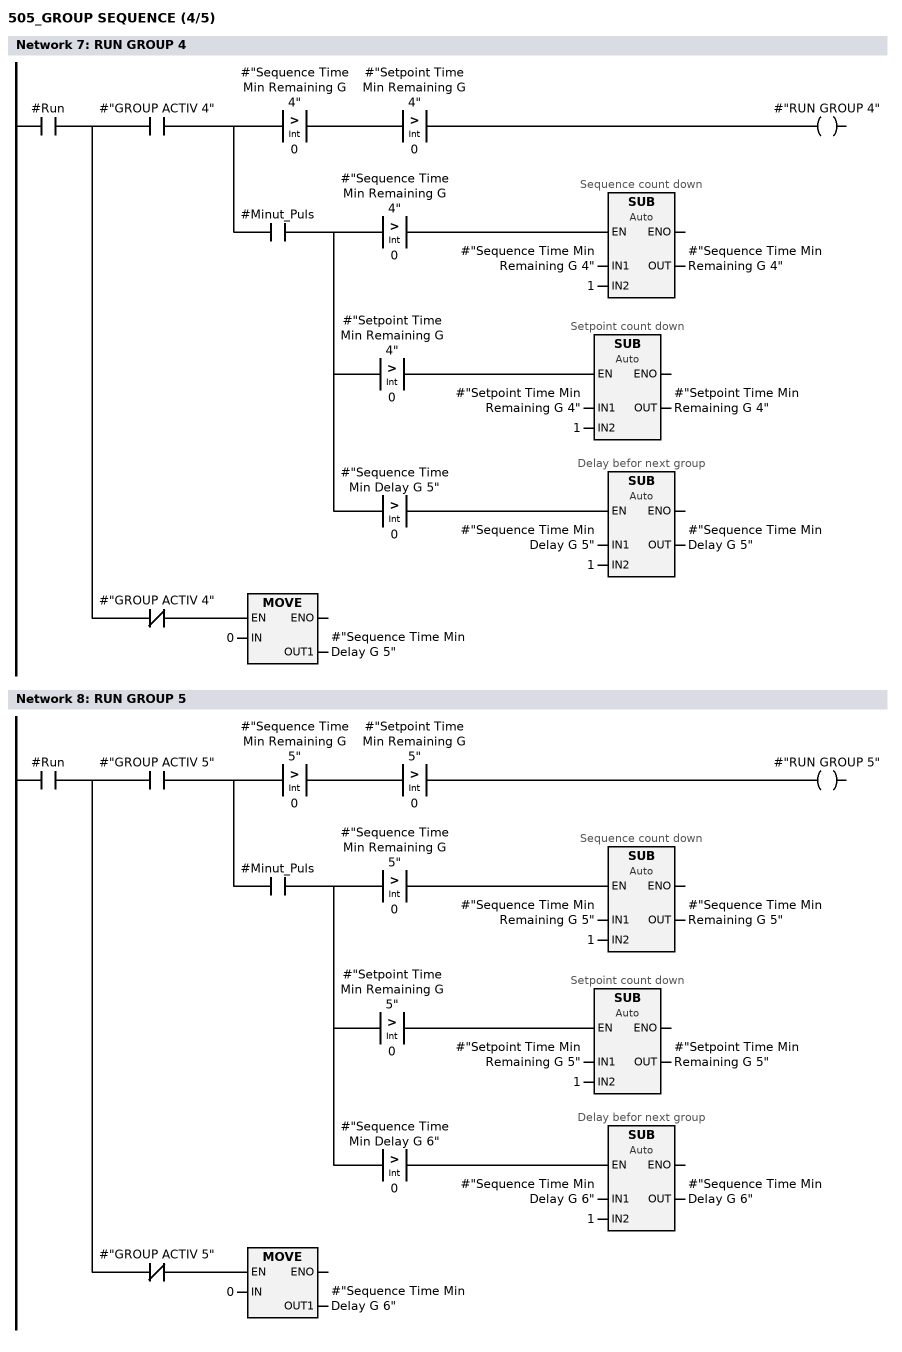
   RUNG wire#powerrail
      Contact( #Run )
      wire#w1
      Contact( #"GROUP ACTIV 4" )
      wire#w2
      { S7_Templates := "SrcType := Int" } GT_Contact(in1 := #"Sequence Time Min Remaining G 4", in2 := 0)
      { S7_Templates := "SrcType := Int" } GT_Contact(in1 := #"Setpoint Time Min Remaining G 4", in2 := 0)
      Coil( #"RUN GROUP 4" )
   END_RUNG
   RUNG wire#w2
      Contact( #Minut_Puls )
      wire#w3
      { S7_Templates := "SrcType := Int" } GT_Contact(in1 := #"Sequence Time Min Remaining G 4", in2 := 0)
      Sub(in1 := #"Sequence Time Min Remaining G 4", in2 := 1, out => #"Sequence Time Min Remaining G 4")   // Sequence count down
   END_RUNG
   RUNG wire#w3
      { S7_Templates := "SrcType := Int" } GT_Contact(in1 := #"Setpoint Time Min Remaining G 4", in2 := 0)
      Sub(in1 := #"Setpoint Time Min Remaining G 4", in2 := 1, out => #"Setpoint Time Min Remaining G 4")   // Setpoint count down
   END_RUNG
   RUNG wire#w3
      { S7_Templates := "SrcType := Int" } GT_Contact(in1 := #"Sequence Time Min Delay G 5", in2 := 0)
      Sub(in1 := #"Sequence Time Min Delay G 5", in2 := 1, out => #"Sequence Time Min Delay G 5")   // Delay befor next group
   END_RUNG
   RUNG wire#w1
      I_Contact( #"GROUP ACTIV 4" )
      Move(in := 0, out1 => #"Sequence Time Min Delay G 5")
   END_RUNG
   // the same network as SCL:
   #_w1 := #Run AND #"GROUP ACTIV 4";
   #"RUN GROUP 4" := #_w1 AND (#"Sequence Time Min Remaining G 4" > 0) AND (#"Setpoint Time Min Remaining G 4" > 0);
   #_w2 := #_w1 AND #Minut_Puls;
   IF #_w2 AND (#"Sequence Time Min Remaining G 4" > 0) THEN
       #"Sequence Time Min Remaining G 4" := #"Sequence Time Min Remaining G 4" - 1;   // Sequence count down
   END_IF;
   IF #_w2 AND (#"Setpoint Time Min Remaining G 4" > 0) THEN
       #"Setpoint Time Min Remaining G 4" := #"Setpoint Time Min Remaining G 4" - 1;   // Setpoint count down
   END_IF;
   IF #_w2 AND (#"Sequence Time Min Delay G 5" > 0) THEN
       #"Sequence Time Min Delay G 5" := #"Sequence Time Min Delay G 5" - 1;   // Delay befor next group
   END_IF;
   IF #Run AND NOT #"GROUP ACTIV 4" THEN #"Sequence Time Min Delay G 5" := 0; END_IF;
END_REGION

REGION Network 8: RUN GROUP 5
   RUNG wire#powerrail
      Contact( #Run )
      wire#w1
      Contact( #"GROUP ACTIV 5" )
      wire#w2
      { S7_Templates := "SrcType := Int" } GT_Contact(in1 := #"Sequence Time Min Remaining G 5", in2 := 0)
      { S7_Templates := "SrcType := Int" } GT_Contact(in1 := #"Setpoint Time Min Remaining G 5", in2 := 0)
      Coil( #"RUN GROUP 5" )
   END_RUNG
   RUNG wire#w2
      Contact( #Minut_Puls )
      wire#w3
      { S7_Templates := "SrcType := Int" } GT_Contact(in1 := #"Sequence Time Min Remaining G 5", in2 := 0)
      Sub(in1 := #"Sequence Time Min Remaining G 5", in2 := 1, out => #"Sequence Time Min Remaining G 5")   // Sequence count down
   END_RUNG
   RUNG wire#w3
      { S7_Templates := "SrcType := Int" } GT_Contact(in1 := #"Setpoint Time Min Remaining G 5", in2 := 0)
      Sub(in1 := #"Setpoint Time Min Remaining G 5", in2 := 1, out => #"Setpoint Time Min Remaining G 5")   // Setpoint count down
   END_RUNG
   RUNG wire#w3
      { S7_Templates := "SrcType := Int" } GT_Contact(in1 := #"Sequence Time Min Delay G 6", in2 := 0)
      Sub(in1 := #"Sequence Time Min Delay G 6", in2 := 1, out => #"Sequence Time Min Delay G 6")   // Delay befor next group
   END_RUNG
   RUNG wire#w1
      I_Contact( #"GROUP ACTIV 5" )
      Move(in := 0, out1 => #"Sequence Time Min Delay G 6")
   END_RUNG
   // the same network as SCL:
   #_w1 := #Run AND #"GROUP ACTIV 5";
   #"RUN GROUP 5" := #_w1 AND (#"Sequence Time Min Remaining G 5" > 0) AND (#"Setpoint Time Min Remaining G 5" > 0);
   #_w2 := #_w1 AND #Minut_Puls;
   IF #_w2 AND (#"Sequence Time Min Remaining G 5" > 0) THEN
       #"Sequence Time Min Remaining G 5" := #"Sequence Time Min Remaining G 5" - 1;   // Sequence count down
   END_IF;
   IF #_w2 AND (#"Setpoint Time Min Remaining G 5" > 0) THEN
       #"Setpoint Time Min Remaining G 5" := #"Setpoint Time Min Remaining G 5" - 1;   // Setpoint count down
   END_IF;
   IF #_w2 AND (#"Sequence Time Min Delay G 6" > 0) THEN
       #"Sequence Time Min Delay G 6" := #"Sequence Time Min Delay G 6" - 1;   // Delay befor next group
   END_IF;
   IF #Run AND NOT #"GROUP ACTIV 5" THEN #"Sequence Time Min Delay G 6" := 0; END_IF;
END_REGION

REGION Network 9: RUN GROUP 6
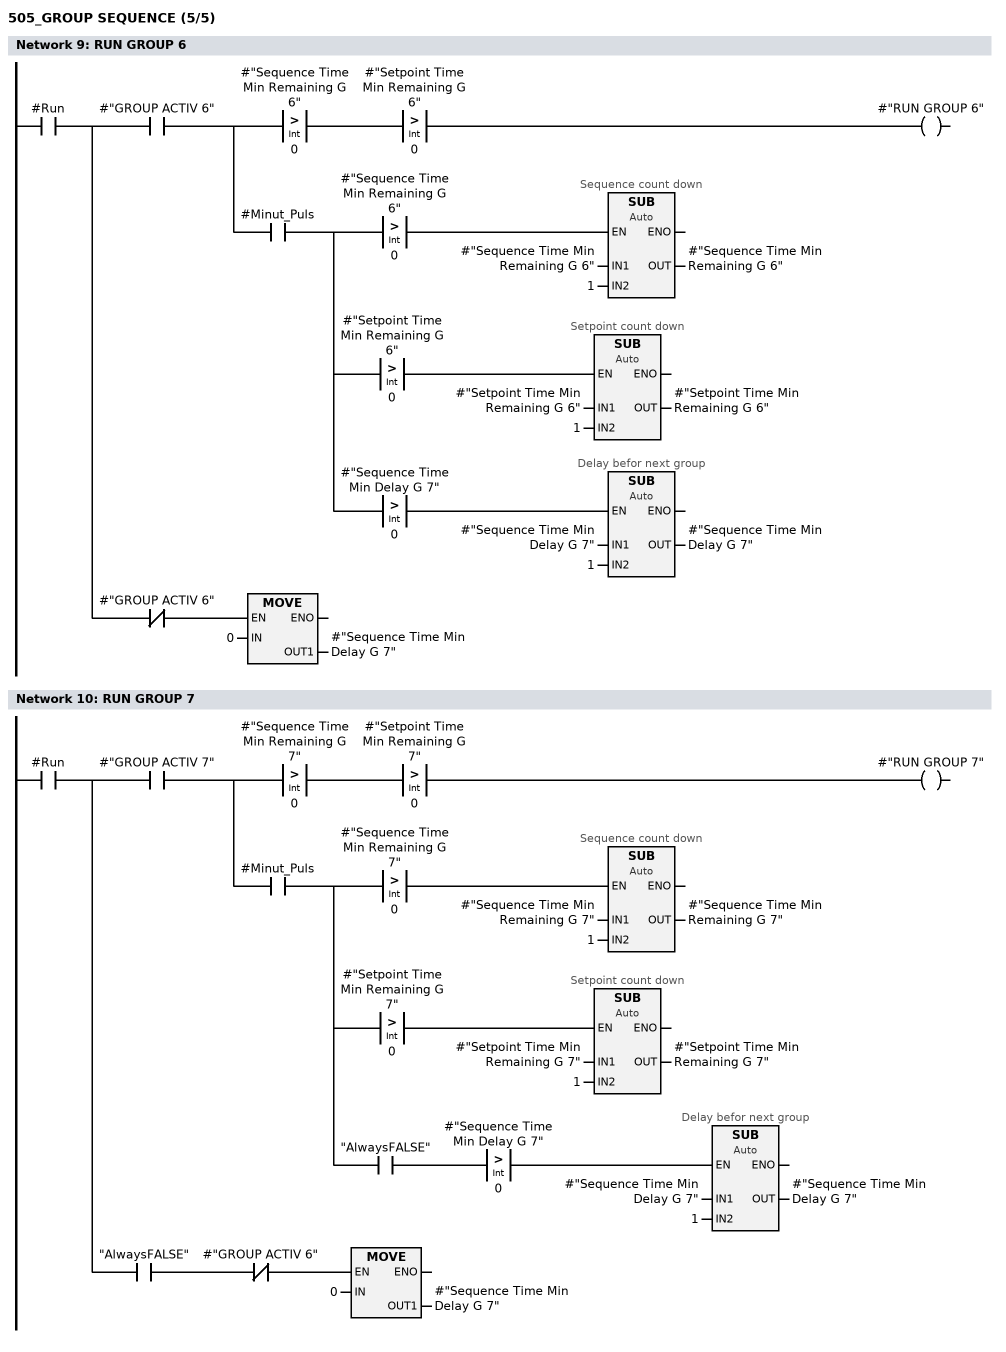
   RUNG wire#powerrail
      Contact( #Run )
      wire#w1
      Contact( #"GROUP ACTIV 6" )
      wire#w2
      { S7_Templates := "SrcType := Int" } GT_Contact(in1 := #"Sequence Time Min Remaining G 6", in2 := 0)
      { S7_Templates := "SrcType := Int" } GT_Contact(in1 := #"Setpoint Time Min Remaining G 6", in2 := 0)
      Coil( #"RUN GROUP 6" )
   END_RUNG
   RUNG wire#w2
      Contact( #Minut_Puls )
      wire#w3
      { S7_Templates := "SrcType := Int" } GT_Contact(in1 := #"Sequence Time Min Remaining G 6", in2 := 0)
      Sub(in1 := #"Sequence Time Min Remaining G 6", in2 := 1, out => #"Sequence Time Min Remaining G 6")   // Sequence count down
   END_RUNG
   RUNG wire#w3
      { S7_Templates := "SrcType := Int" } GT_Contact(in1 := #"Setpoint Time Min Remaining G 6", in2 := 0)
      Sub(in1 := #"Setpoint Time Min Remaining G 6", in2 := 1, out => #"Setpoint Time Min Remaining G 6")   // Setpoint count down
   END_RUNG
   RUNG wire#w3
      { S7_Templates := "SrcType := Int" } GT_Contact(in1 := #"Sequence Time Min Delay G 7", in2 := 0)
      Sub(in1 := #"Sequence Time Min Delay G 7", in2 := 1, out => #"Sequence Time Min Delay G 7")   // Delay befor next group
   END_RUNG
   RUNG wire#w1
      I_Contact( #"GROUP ACTIV 6" )
      Move(in := 0, out1 => #"Sequence Time Min Delay G 7")
   END_RUNG
   // the same network as SCL:
   #_w1 := #Run AND #"GROUP ACTIV 6";
   #"RUN GROUP 6" := #_w1 AND (#"Sequence Time Min Remaining G 6" > 0) AND (#"Setpoint Time Min Remaining G 6" > 0);
   #_w2 := #_w1 AND #Minut_Puls;
   IF #_w2 AND (#"Sequence Time Min Remaining G 6" > 0) THEN
       #"Sequence Time Min Remaining G 6" := #"Sequence Time Min Remaining G 6" - 1;   // Sequence count down
   END_IF;
   IF #_w2 AND (#"Setpoint Time Min Remaining G 6" > 0) THEN
       #"Setpoint Time Min Remaining G 6" := #"Setpoint Time Min Remaining G 6" - 1;   // Setpoint count down
   END_IF;
   IF #_w2 AND (#"Sequence Time Min Delay G 7" > 0) THEN
       #"Sequence Time Min Delay G 7" := #"Sequence Time Min Delay G 7" - 1;   // Delay befor next group
   END_IF;
   IF #Run AND NOT #"GROUP ACTIV 6" THEN #"Sequence Time Min Delay G 7" := 0; END_IF;
END_REGION

REGION Network 10: RUN GROUP 7
   RUNG wire#powerrail
      Contact( #Run )
      wire#w1
      Contact( #"GROUP ACTIV 7" )
      wire#w2
      { S7_Templates := "SrcType := Int" } GT_Contact(in1 := #"Sequence Time Min Remaining G 7", in2 := 0)
      { S7_Templates := "SrcType := Int" } GT_Contact(in1 := #"Setpoint Time Min Remaining G 7", in2 := 0)
      Coil( #"RUN GROUP 7" )
   END_RUNG
   RUNG wire#w2
      Contact( #Minut_Puls )
      wire#w3
      { S7_Templates := "SrcType := Int" } GT_Contact(in1 := #"Sequence Time Min Remaining G 7", in2 := 0)
      Sub(in1 := #"Sequence Time Min Remaining G 7", in2 := 1, out => #"Sequence Time Min Remaining G 7")   // Sequence count down
   END_RUNG
   RUNG wire#w3
      { S7_Templates := "SrcType := Int" } GT_Contact(in1 := #"Setpoint Time Min Remaining G 7", in2 := 0)
      Sub(in1 := #"Setpoint Time Min Remaining G 7", in2 := 1, out => #"Setpoint Time Min Remaining G 7")   // Setpoint count down
   END_RUNG
   RUNG wire#w3
      Contact( "AlwaysFALSE" )
      { S7_Templates := "SrcType := Int" } GT_Contact(in1 := #"Sequence Time Min Delay G 7", in2 := 0)
      Sub(in1 := #"Sequence Time Min Delay G 7", in2 := 1, out => #"Sequence Time Min Delay G 7")   // Delay befor next group
   END_RUNG
   RUNG wire#w1
      Contact( "AlwaysFALSE" )
      I_Contact( #"GROUP ACTIV 6" )
      Move(in := 0, out1 => #"Sequence Time Min Delay G 7")
   END_RUNG
   // the same network as SCL:
   #_w1 := #Run AND #"GROUP ACTIV 7";
   #"RUN GROUP 7" := #_w1 AND (#"Sequence Time Min Remaining G 7" > 0) AND (#"Setpoint Time Min Remaining G 7" > 0);
   #_w2 := #_w1 AND #Minut_Puls;
   IF #_w2 AND (#"Sequence Time Min Remaining G 7" > 0) THEN
       #"Sequence Time Min Remaining G 7" := #"Sequence Time Min Remaining G 7" - 1;   // Sequence count down
   END_IF;
   IF #_w2 AND (#"Setpoint Time Min Remaining G 7" > 0) THEN
       #"Setpoint Time Min Remaining G 7" := #"Setpoint Time Min Remaining G 7" - 1;   // Setpoint count down
   END_IF;
   IF #_w2 AND "AlwaysFALSE" AND (#"Sequence Time Min Delay G 7" > 0) THEN
       #"Sequence Time Min Delay G 7" := #"Sequence Time Min Delay G 7" - 1;   // Delay befor next group
   END_IF;
   IF #Run AND "AlwaysFALSE" AND NOT #"GROUP ACTIV 6" THEN #"Sequence Time Min Delay G 7" := 0; END_IF;
END_REGION
END_FUNCTION_BLOCK

FUNCTION_BLOCK "Binary Imputs ADD"   // FB506, LAD
{ S7_Optimized_Access := 'TRUE' }
VERSION : 0.1
   VAR_INPUT
      "BI 1" : Bool;
      "BI 2" : Bool;
      "BI 3" : Bool;
      "BI 4" : Bool;
      "BI 5" : Bool;
      "BI 6" : Bool;
      "BI 7" : Bool;
      "BI 8" : Bool;
      "BI 9" : Bool;
      "BI 10" : Bool;
      "BI 11" : Bool;
      "BI 12" : Bool;
      "BI 13" : Bool;
      "BI 14" : Bool;
      "BI 15" : Bool;
      "BI 16" : Bool;
      "BI 17" : Bool;
      "BI 18" : Bool;
      "BI 19" : Bool;
      "BI 20" : Bool;
      "BI 21" : Bool;
      "BI 22" : Bool;
      "BI 23" : Bool;
      "BI 24" : Bool;
   END_VAR
   VAR_OUTPUT
      "BI Number" : Int;
   END_VAR
   VAR
      "BI Interm 1" : Int;
      "BI Interm 2" : Int;
      "BI Interm 3" : Int;
      "BI Interm 4" : Int;
      "BI Interm 5" : Int;
      "BI Interm 6" : Int;
      "BI Interm 7" : Int;
      "BI Interm 8" : Int;
      "BI Interm 9" : Int;
      "BI Interm 10" : Int;
      "BI Interm 11" : Int;
      "BI Interm 12" : Int;
      "BI Interm 13" : Int;
      "BI Interm 14" : Int;
      "BI Interm 15" : Int;
      "BI Interm 16" : Int;
      "BI Interm 17" : Int;
      "BI Interm 18" : Int;
      "BI Interm 19" : Int;
      "BI Interm 20" : Int;
      "BI Interm 21" : Int;
      "BI Interm 22" : Int;
      "BI Interm 23" : Int;
      "BI Interm 24" : Int;
   END_VAR
BEGIN

REGION Network 1: 1
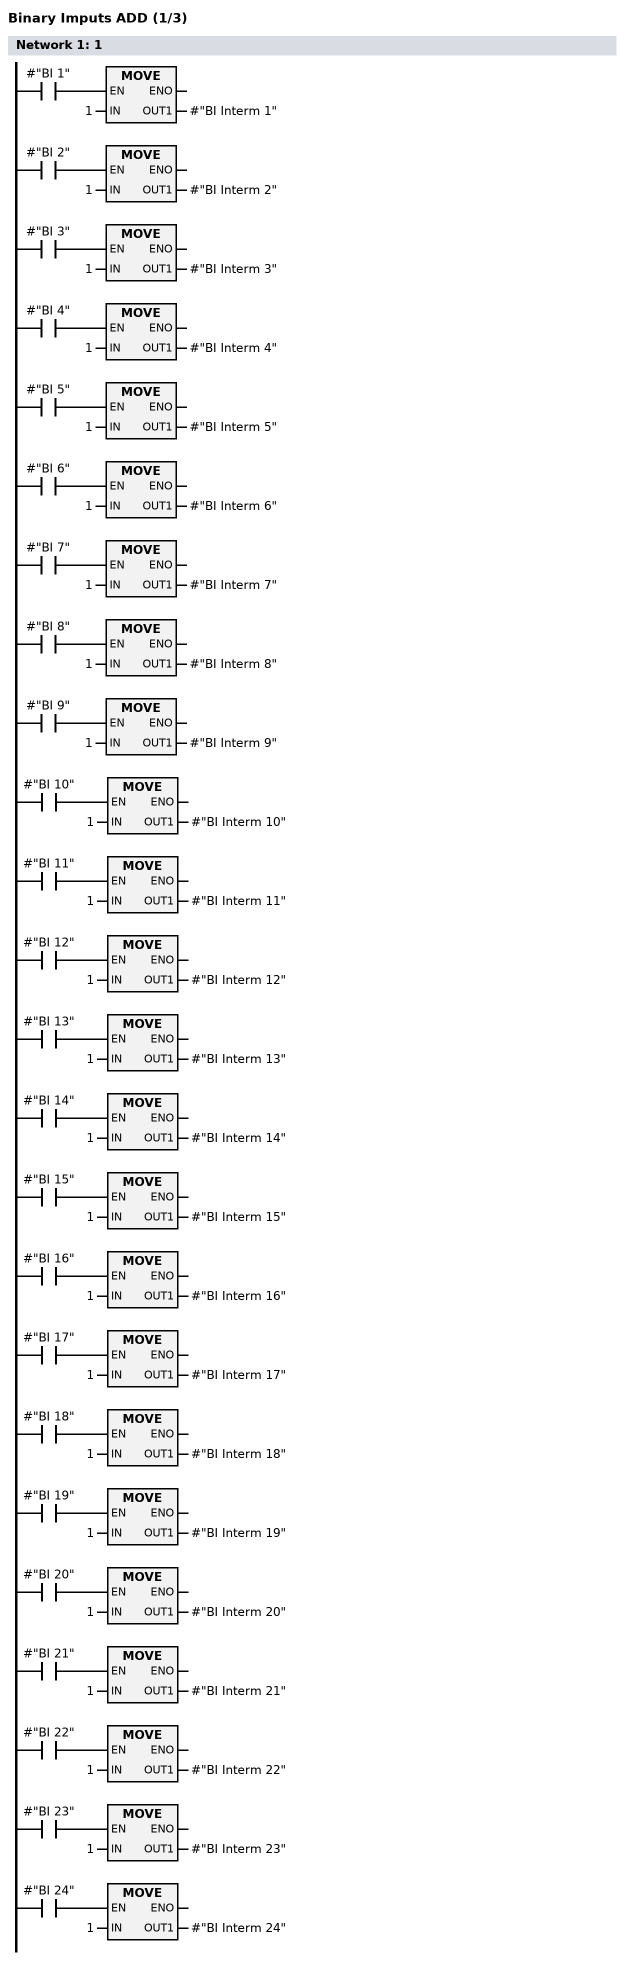
   RUNG wire#powerrail
      Contact( #"BI 1" )
      Move(in := 1, out1 => #"BI Interm 1")
   END_RUNG
   RUNG wire#powerrail
      Contact( #"BI 2" )
      Move(in := 1, out1 => #"BI Interm 2")
   END_RUNG
   RUNG wire#powerrail
      Contact( #"BI 3" )
      Move(in := 1, out1 => #"BI Interm 3")
   END_RUNG
   RUNG wire#powerrail
      Contact( #"BI 4" )
      Move(in := 1, out1 => #"BI Interm 4")
   END_RUNG
   RUNG wire#powerrail
      Contact( #"BI 5" )
      Move(in := 1, out1 => #"BI Interm 5")
   END_RUNG
   RUNG wire#powerrail
      Contact( #"BI 6" )
      Move(in := 1, out1 => #"BI Interm 6")
   END_RUNG
   RUNG wire#powerrail
      Contact( #"BI 7" )
      Move(in := 1, out1 => #"BI Interm 7")
   END_RUNG
   RUNG wire#powerrail
      Contact( #"BI 8" )
      Move(in := 1, out1 => #"BI Interm 8")
   END_RUNG
   RUNG wire#powerrail
      Contact( #"BI 9" )
      Move(in := 1, out1 => #"BI Interm 9")
   END_RUNG
   RUNG wire#powerrail
      Contact( #"BI 10" )
      Move(in := 1, out1 => #"BI Interm 10")
   END_RUNG
   RUNG wire#powerrail
      Contact( #"BI 11" )
      Move(in := 1, out1 => #"BI Interm 11")
   END_RUNG
   RUNG wire#powerrail
      Contact( #"BI 12" )
      Move(in := 1, out1 => #"BI Interm 12")
   END_RUNG
   RUNG wire#powerrail
      Contact( #"BI 13" )
      Move(in := 1, out1 => #"BI Interm 13")
   END_RUNG
   RUNG wire#powerrail
      Contact( #"BI 14" )
      Move(in := 1, out1 => #"BI Interm 14")
   END_RUNG
   RUNG wire#powerrail
      Contact( #"BI 15" )
      Move(in := 1, out1 => #"BI Interm 15")
   END_RUNG
   RUNG wire#powerrail
      Contact( #"BI 16" )
      Move(in := 1, out1 => #"BI Interm 16")
   END_RUNG
   RUNG wire#powerrail
      Contact( #"BI 17" )
      Move(in := 1, out1 => #"BI Interm 17")
   END_RUNG
   RUNG wire#powerrail
      Contact( #"BI 18" )
      Move(in := 1, out1 => #"BI Interm 18")
   END_RUNG
   RUNG wire#powerrail
      Contact( #"BI 19" )
      Move(in := 1, out1 => #"BI Interm 19")
   END_RUNG
   RUNG wire#powerrail
      Contact( #"BI 20" )
      Move(in := 1, out1 => #"BI Interm 20")
   END_RUNG
   RUNG wire#powerrail
      Contact( #"BI 21" )
      Move(in := 1, out1 => #"BI Interm 21")
   END_RUNG
   RUNG wire#powerrail
      Contact( #"BI 22" )
      Move(in := 1, out1 => #"BI Interm 22")
   END_RUNG
   RUNG wire#powerrail
      Contact( #"BI 23" )
      Move(in := 1, out1 => #"BI Interm 23")
   END_RUNG
   RUNG wire#powerrail
      Contact( #"BI 24" )
      Move(in := 1, out1 => #"BI Interm 24")
   END_RUNG
   // the same network as SCL:
   IF #"BI 1" THEN #"BI Interm 1" := 1; END_IF;
   IF #"BI 2" THEN #"BI Interm 2" := 1; END_IF;
   IF #"BI 3" THEN #"BI Interm 3" := 1; END_IF;
   IF #"BI 4" THEN #"BI Interm 4" := 1; END_IF;
   IF #"BI 5" THEN #"BI Interm 5" := 1; END_IF;
   IF #"BI 6" THEN #"BI Interm 6" := 1; END_IF;
   IF #"BI 7" THEN #"BI Interm 7" := 1; END_IF;
   IF #"BI 8" THEN #"BI Interm 8" := 1; END_IF;
   IF #"BI 9" THEN #"BI Interm 9" := 1; END_IF;
   IF #"BI 10" THEN #"BI Interm 10" := 1; END_IF;
   IF #"BI 11" THEN #"BI Interm 11" := 1; END_IF;
   IF #"BI 12" THEN #"BI Interm 12" := 1; END_IF;
   IF #"BI 13" THEN #"BI Interm 13" := 1; END_IF;
   IF #"BI 14" THEN #"BI Interm 14" := 1; END_IF;
   IF #"BI 15" THEN #"BI Interm 15" := 1; END_IF;
   IF #"BI 16" THEN #"BI Interm 16" := 1; END_IF;
   IF #"BI 17" THEN #"BI Interm 17" := 1; END_IF;
   IF #"BI 18" THEN #"BI Interm 18" := 1; END_IF;
   IF #"BI 19" THEN #"BI Interm 19" := 1; END_IF;
   IF #"BI 20" THEN #"BI Interm 20" := 1; END_IF;
   IF #"BI 21" THEN #"BI Interm 21" := 1; END_IF;
   IF #"BI 22" THEN #"BI Interm 22" := 1; END_IF;
   IF #"BI 23" THEN #"BI Interm 23" := 1; END_IF;
   IF #"BI 24" THEN #"BI Interm 24" := 1; END_IF;
END_REGION

REGION Network 2: 0
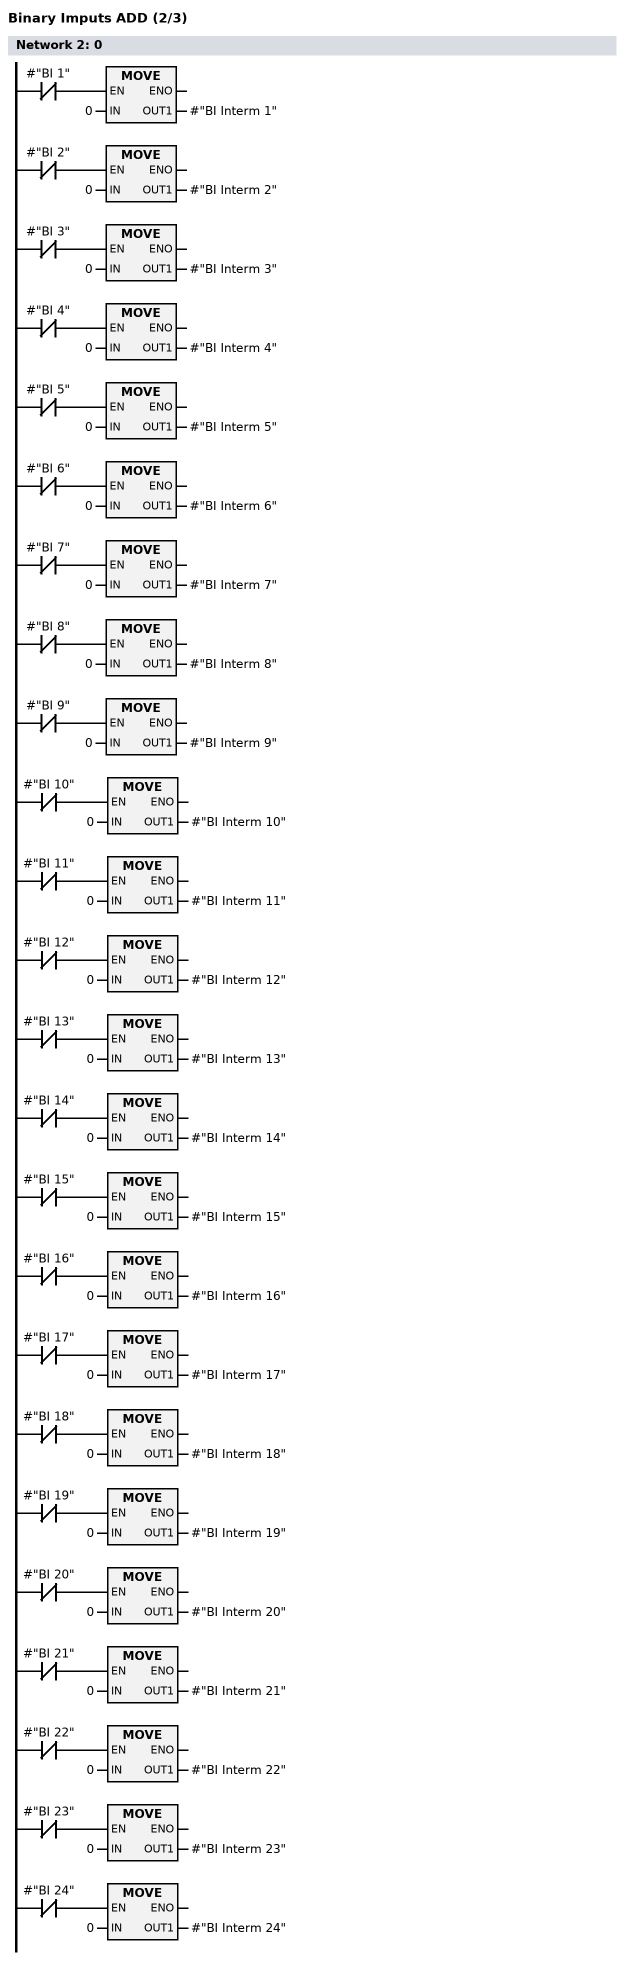
   RUNG wire#powerrail
      I_Contact( #"BI 1" )
      Move(in := 0, out1 => #"BI Interm 1")
   END_RUNG
   RUNG wire#powerrail
      I_Contact( #"BI 2" )
      Move(in := 0, out1 => #"BI Interm 2")
   END_RUNG
   RUNG wire#powerrail
      I_Contact( #"BI 3" )
      Move(in := 0, out1 => #"BI Interm 3")
   END_RUNG
   RUNG wire#powerrail
      I_Contact( #"BI 4" )
      Move(in := 0, out1 => #"BI Interm 4")
   END_RUNG
   RUNG wire#powerrail
      I_Contact( #"BI 5" )
      Move(in := 0, out1 => #"BI Interm 5")
   END_RUNG
   RUNG wire#powerrail
      I_Contact( #"BI 6" )
      Move(in := 0, out1 => #"BI Interm 6")
   END_RUNG
   RUNG wire#powerrail
      I_Contact( #"BI 7" )
      Move(in := 0, out1 => #"BI Interm 7")
   END_RUNG
   RUNG wire#powerrail
      I_Contact( #"BI 8" )
      Move(in := 0, out1 => #"BI Interm 8")
   END_RUNG
   RUNG wire#powerrail
      I_Contact( #"BI 9" )
      Move(in := 0, out1 => #"BI Interm 9")
   END_RUNG
   RUNG wire#powerrail
      I_Contact( #"BI 10" )
      Move(in := 0, out1 => #"BI Interm 10")
   END_RUNG
   RUNG wire#powerrail
      I_Contact( #"BI 11" )
      Move(in := 0, out1 => #"BI Interm 11")
   END_RUNG
   RUNG wire#powerrail
      I_Contact( #"BI 12" )
      Move(in := 0, out1 => #"BI Interm 12")
   END_RUNG
   RUNG wire#powerrail
      I_Contact( #"BI 13" )
      Move(in := 0, out1 => #"BI Interm 13")
   END_RUNG
   RUNG wire#powerrail
      I_Contact( #"BI 14" )
      Move(in := 0, out1 => #"BI Interm 14")
   END_RUNG
   RUNG wire#powerrail
      I_Contact( #"BI 15" )
      Move(in := 0, out1 => #"BI Interm 15")
   END_RUNG
   RUNG wire#powerrail
      I_Contact( #"BI 16" )
      Move(in := 0, out1 => #"BI Interm 16")
   END_RUNG
   RUNG wire#powerrail
      I_Contact( #"BI 17" )
      Move(in := 0, out1 => #"BI Interm 17")
   END_RUNG
   RUNG wire#powerrail
      I_Contact( #"BI 18" )
      Move(in := 0, out1 => #"BI Interm 18")
   END_RUNG
   RUNG wire#powerrail
      I_Contact( #"BI 19" )
      Move(in := 0, out1 => #"BI Interm 19")
   END_RUNG
   RUNG wire#powerrail
      I_Contact( #"BI 20" )
      Move(in := 0, out1 => #"BI Interm 20")
   END_RUNG
   RUNG wire#powerrail
      I_Contact( #"BI 21" )
      Move(in := 0, out1 => #"BI Interm 21")
   END_RUNG
   RUNG wire#powerrail
      I_Contact( #"BI 22" )
      Move(in := 0, out1 => #"BI Interm 22")
   END_RUNG
   RUNG wire#powerrail
      I_Contact( #"BI 23" )
      Move(in := 0, out1 => #"BI Interm 23")
   END_RUNG
   RUNG wire#powerrail
      I_Contact( #"BI 24" )
      Move(in := 0, out1 => #"BI Interm 24")
   END_RUNG
   // the same network as SCL:
   IF NOT #"BI 1" THEN #"BI Interm 1" := 0; END_IF;
   IF NOT #"BI 2" THEN #"BI Interm 2" := 0; END_IF;
   IF NOT #"BI 3" THEN #"BI Interm 3" := 0; END_IF;
   IF NOT #"BI 4" THEN #"BI Interm 4" := 0; END_IF;
   IF NOT #"BI 5" THEN #"BI Interm 5" := 0; END_IF;
   IF NOT #"BI 6" THEN #"BI Interm 6" := 0; END_IF;
   IF NOT #"BI 7" THEN #"BI Interm 7" := 0; END_IF;
   IF NOT #"BI 8" THEN #"BI Interm 8" := 0; END_IF;
   IF NOT #"BI 9" THEN #"BI Interm 9" := 0; END_IF;
   IF NOT #"BI 10" THEN #"BI Interm 10" := 0; END_IF;
   IF NOT #"BI 11" THEN #"BI Interm 11" := 0; END_IF;
   IF NOT #"BI 12" THEN #"BI Interm 12" := 0; END_IF;
   IF NOT #"BI 13" THEN #"BI Interm 13" := 0; END_IF;
   IF NOT #"BI 14" THEN #"BI Interm 14" := 0; END_IF;
   IF NOT #"BI 15" THEN #"BI Interm 15" := 0; END_IF;
   IF NOT #"BI 16" THEN #"BI Interm 16" := 0; END_IF;
   IF NOT #"BI 17" THEN #"BI Interm 17" := 0; END_IF;
   IF NOT #"BI 18" THEN #"BI Interm 18" := 0; END_IF;
   IF NOT #"BI 19" THEN #"BI Interm 19" := 0; END_IF;
   IF NOT #"BI 20" THEN #"BI Interm 20" := 0; END_IF;
   IF NOT #"BI 21" THEN #"BI Interm 21" := 0; END_IF;
   IF NOT #"BI 22" THEN #"BI Interm 22" := 0; END_IF;
   IF NOT #"BI 23" THEN #"BI Interm 23" := 0; END_IF;
   IF NOT #"BI 24" THEN #"BI Interm 24" := 0; END_IF;
END_REGION

REGION Network 3: ADD
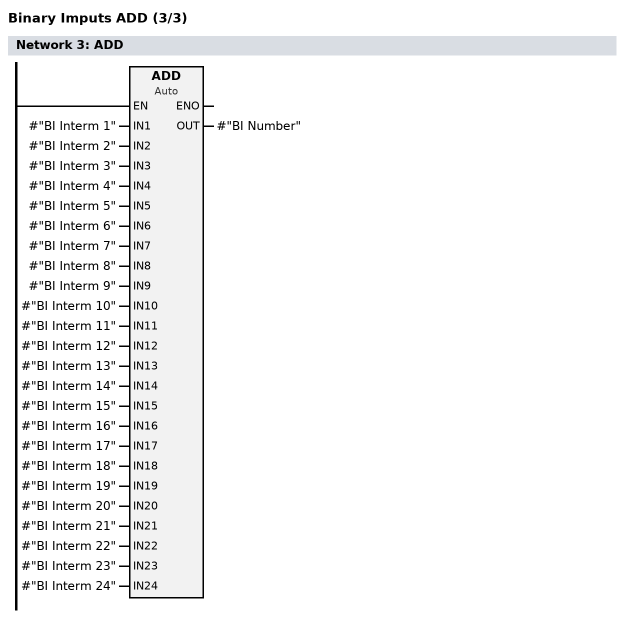
   RUNG wire#powerrail
      Add(in1 := #"BI Interm 1", in2 := #"BI Interm 2", in3 := #"BI Interm 3", in4 := #"BI Interm 4", in5 := #"BI Interm 5", in6 := #"BI Interm 6", in7 := #"BI Interm 7", in8 := #"BI Interm 8", in9 := #"BI Interm 9", in10 := #"BI Interm 10", in11 := #"BI Interm 11", in12 := #"BI Interm 12", in13 := #"BI Interm 13", in14 := #"BI Interm 14", in15 := #"BI Interm 15", in16 := #"BI Interm 16", in17 := #"BI Interm 17", in18 := #"BI Interm 18", in19 := #"BI Interm 19", in20 := #"BI Interm 20", in21 := #"BI Interm 21", in22 := #"BI Interm 22", in23 := #"BI Interm 23", in24 := #"BI Interm 24", out => #"BI Number")
   END_RUNG
   // the same network as SCL:
   #"BI Number" := #"BI Interm 1" + #"BI Interm 2" + #"BI Interm 3" + #"BI Interm 4" + #"BI Interm 5" + #"BI Interm 6" + #"BI Interm 7" + #"BI Interm 8" + #"BI Interm 9" + #"BI Interm 10" + #"BI Interm 11" + #"BI Interm 12" + #"BI Interm 13" + #"BI Interm 14" + #"BI Interm 15" + #"BI Interm 16" + #"BI Interm 17" + #"BI Interm 18" + #"BI Interm 19" + #"BI Interm 20" + #"BI Interm 21" + #"BI Interm 22" + #"BI Interm 23" + #"BI Interm 24";
END_REGION
END_FUNCTION_BLOCK

FUNCTION_BLOCK "HMI Indication Logic"   // FB507, LAD
{ S7_Optimized_Access := 'TRUE' }
VERSION : 0.1
   VAR_OUTPUT
      "FA Mode Selected" : Bool;
      "Tank Selected" : Bool;
      "Sequence Finished" : Bool;
   END_VAR
   VAR
      IEC_Timer_0_Instance : TON_TIME;
   END_VAR
BEGIN

REGION Network 1: FA Mode Selected
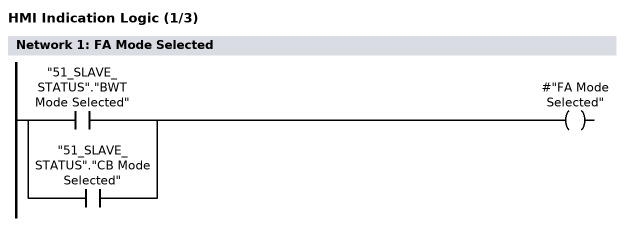
   RUNG wire#powerrail
      Contact( "51_SLAVE_STATUS"."BWT Mode Selected" )
      wire#w1
      Coil( #"FA Mode Selected" )
   END_RUNG
   RUNG wire#powerrail
      Contact( "51_SLAVE_STATUS"."CB Mode Selected" )
   END_RUNG wire#w1
   // the same network as SCL:
   #"FA Mode Selected" := "51_SLAVE_STATUS"."BWT Mode Selected" OR "51_SLAVE_STATUS"."CB Mode Selected";
END_REGION

REGION Network 2: Tank Selected
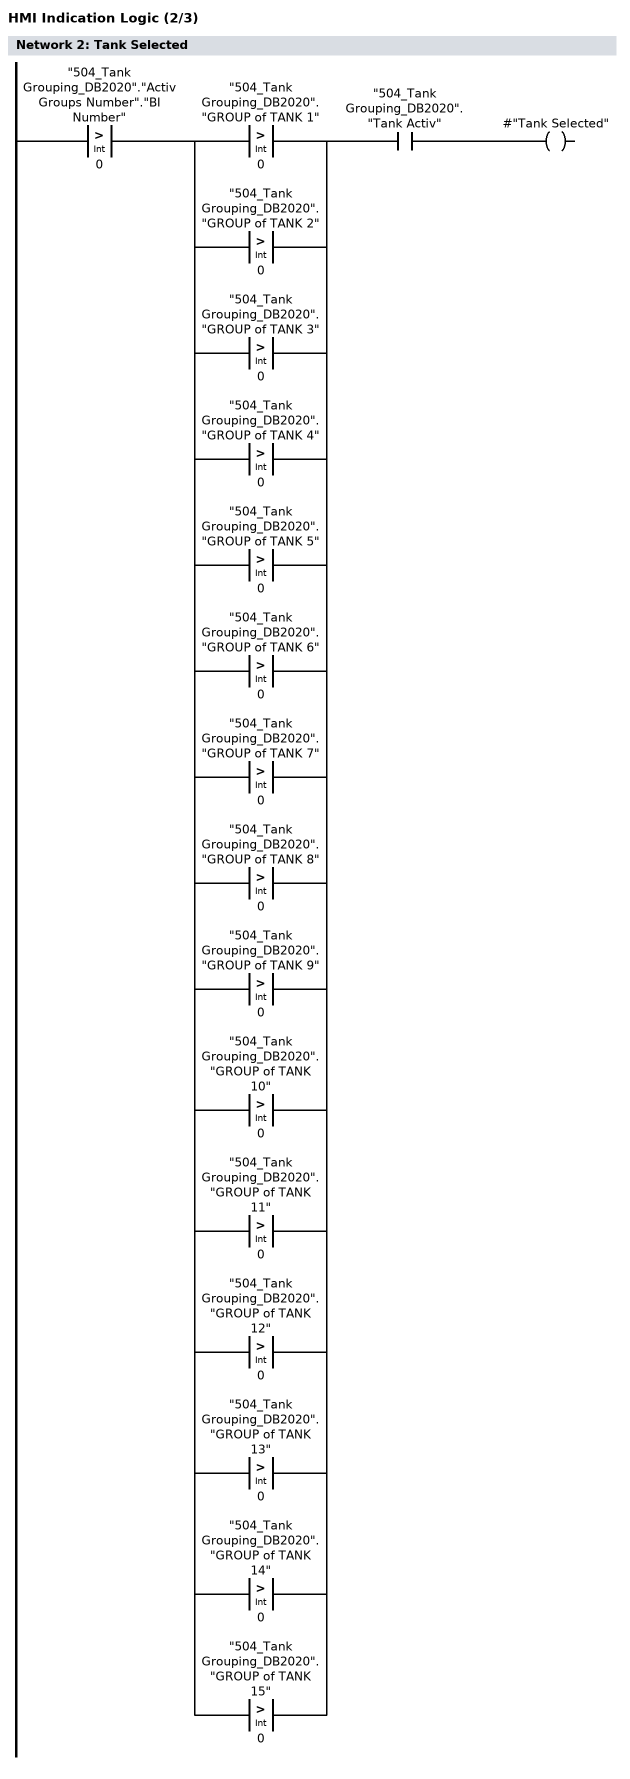
   RUNG wire#powerrail
      { S7_Templates := "SrcType := Int" } GT_Contact(in1 := "504_Tank Grouping_DB2020"."Activ Groups Number"."BI Number", in2 := 0)
      wire#w1
      { S7_Templates := "SrcType := Int" } GT_Contact(in1 := "504_Tank Grouping_DB2020"."GROUP of TANK 1", in2 := 0)
      wire#w2
      Contact( "504_Tank Grouping_DB2020"."Tank Activ" )
      Coil( #"Tank Selected" )
   END_RUNG
   RUNG wire#w1
      { S7_Templates := "SrcType := Int" } GT_Contact(in1 := "504_Tank Grouping_DB2020"."GROUP of TANK 2", in2 := 0)
   END_RUNG wire#w2
   RUNG wire#w1
      { S7_Templates := "SrcType := Int" } GT_Contact(in1 := "504_Tank Grouping_DB2020"."GROUP of TANK 3", in2 := 0)
   END_RUNG wire#w2
   RUNG wire#w1
      { S7_Templates := "SrcType := Int" } GT_Contact(in1 := "504_Tank Grouping_DB2020"."GROUP of TANK 4", in2 := 0)
   END_RUNG wire#w2
   RUNG wire#w1
      { S7_Templates := "SrcType := Int" } GT_Contact(in1 := "504_Tank Grouping_DB2020"."GROUP of TANK 5", in2 := 0)
   END_RUNG wire#w2
   RUNG wire#w1
      { S7_Templates := "SrcType := Int" } GT_Contact(in1 := "504_Tank Grouping_DB2020"."GROUP of TANK 6", in2 := 0)
   END_RUNG wire#w2
   RUNG wire#w1
      { S7_Templates := "SrcType := Int" } GT_Contact(in1 := "504_Tank Grouping_DB2020"."GROUP of TANK 7", in2 := 0)
   END_RUNG wire#w2
   RUNG wire#w1
      { S7_Templates := "SrcType := Int" } GT_Contact(in1 := "504_Tank Grouping_DB2020"."GROUP of TANK 8", in2 := 0)
   END_RUNG wire#w2
   RUNG wire#w1
      { S7_Templates := "SrcType := Int" } GT_Contact(in1 := "504_Tank Grouping_DB2020"."GROUP of TANK 9", in2 := 0)
   END_RUNG wire#w2
   RUNG wire#w1
      { S7_Templates := "SrcType := Int" } GT_Contact(in1 := "504_Tank Grouping_DB2020"."GROUP of TANK 10", in2 := 0)
   END_RUNG wire#w2
   RUNG wire#w1
      { S7_Templates := "SrcType := Int" } GT_Contact(in1 := "504_Tank Grouping_DB2020"."GROUP of TANK 11", in2 := 0)
   END_RUNG wire#w2
   RUNG wire#w1
      { S7_Templates := "SrcType := Int" } GT_Contact(in1 := "504_Tank Grouping_DB2020"."GROUP of TANK 12", in2 := 0)
   END_RUNG wire#w2
   RUNG wire#w1
      { S7_Templates := "SrcType := Int" } GT_Contact(in1 := "504_Tank Grouping_DB2020"."GROUP of TANK 13", in2 := 0)
   END_RUNG wire#w2
   RUNG wire#w1
      { S7_Templates := "SrcType := Int" } GT_Contact(in1 := "504_Tank Grouping_DB2020"."GROUP of TANK 14", in2 := 0)
   END_RUNG wire#w2
   RUNG wire#w1
      { S7_Templates := "SrcType := Int" } GT_Contact(in1 := "504_Tank Grouping_DB2020"."GROUP of TANK 15", in2 := 0)
   END_RUNG wire#w2
   // the same network as SCL:
   #"Tank Selected" := ("504_Tank Grouping_DB2020"."Activ Groups Number"."BI Number" > 0) AND (("504_Tank Grouping_DB2020"."GROUP of TANK 1" > 0) OR ("504_Tank Grouping_DB2020"."GROUP of TANK 2" > 0) OR ("504_Tank Grouping_DB2020"."GROUP of TANK 3" > 0) OR ("504_Tank Grouping_DB2020"."GROUP of TANK 4" > 0) OR ("504_Tank Grouping_DB2020"."GROUP of TANK 5" > 0) OR ("504_Tank Grouping_DB2020"."GROUP of TANK 6" > 0) OR ("504_Tank Grouping_DB2020"."GROUP of TANK 7" > 0) OR ("504_Tank Grouping_DB2020"."GROUP of TANK 8" > 0) OR ("504_Tank Grouping_DB2020"."GROUP of TANK 9" > 0) OR ("504_Tank Grouping_DB2020"."GROUP of TANK 10" > 0) OR ("504_Tank Grouping_DB2020"."GROUP of TANK 11" > 0) OR ("504_Tank Grouping_DB2020"."GROUP of TANK 12" > 0) OR ("504_Tank Grouping_DB2020"."GROUP of TANK 13" > 0) OR ("504_Tank Grouping_DB2020"."GROUP of TANK 14" > 0) OR ("504_Tank Grouping_DB2020"."GROUP of TANK 15" > 0)) AND "504_Tank Grouping_DB2020"."Tank Activ";
END_REGION

REGION Network 3: Sequence finished
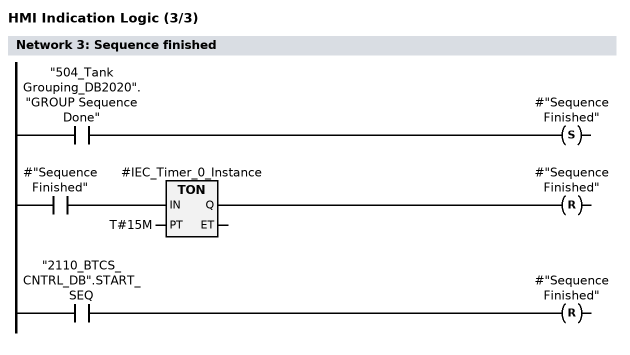
   IF "504_Tank Grouping_DB2020"."GROUP Sequence Done" THEN #"Sequence Finished" := TRUE; END_IF;
   #IEC_Timer_0_Instance(IN := #"Sequence Finished", PT := T#15M);   // TON
   IF #IEC_Timer_0_Instance.Q THEN #"Sequence Finished" := FALSE; END_IF;
   IF "2110_BTCS_CNTRL_DB".START_SEQ THEN #"Sequence Finished" := FALSE; END_IF;
END_REGION
END_FUNCTION_BLOCK

FUNCTION_BLOCK "503_ALARM CHCK"   // FB508, LAD
{ S7_Optimized_Access := 'TRUE' }
VERSION : 0.1
   VAR_INPUT
      "Alarm Word 1" : Word;
      "Alarm Word 2" : Word;
      "Alarm Word 3" : Word;
      "Alarm Word 4" : Word;
      "Alarm Word 5" : Word;
      "Alarm Word 6" : Word;
      "Alarm Word 7" : Word;
      "Alarm Word 8" : Word;
      "Alarm Word 9" : Word;
      "Alarm Word 10" : Word;
      "Alarm Word 11" : Word;
      "Alarm Word 12" : Word;
      "Alarm Word 13" : Word;
      "Alarm Word 14" : Word;
      "Alarm Word 15" : Word;
      "Alarm Word 16" : Word;
      "Reset Alarm" : Bool;
   END_VAR
   VAR_OUTPUT
      "Sound Alarm" : Bool;
   END_VAR
   VAR
      "Alarm Word Interm 1" : Word;
      "Alarm Word Interm 2" : Word;
      "Alarm Word Interm 3" : Word;
      "Alarm Word Interm 4" : Word;
      "Alarm Word Interm 5" : Word;
      "Alarm Word Interm 6" : Word;
      "Alarm Word Interm 7" : Word;
      "Alarm Word Interm 8" : Word;
      "Alarm Word Interm 9" : Word;
      "Alarm Word Interm 10" : Word;
      "Alarm Word Interm 11" : Word;
      "Alarm Word Interm 12" : Word;
      "Alarm Word Interm 13" : Word;
      "Alarm Word Interm 14" : Word;
      "Alarm Word Interm 15" : Word;
      "Alarm Word Interm 16" : Word;
      "Alarm Word bool 1" : Bool;
      "Alarm Word bool 2" : Bool;
      "Alarm Word bool 3" : Bool;
      "Alarm Word bool 4" : Bool;
      "Alarm Word bool 5" : Bool;
      "Alarm Word bool 6" : Bool;
      "Alarm Word bool 7" : Bool;
      "Alarm Word bool 8" : Bool;
      "Alarm Word bool 9" : Bool;
      "Alarm Word bool 10" : Bool;
      "Alarm Word bool 11" : Bool;
      "Alarm Word bool 12" : Bool;
      "Alarm Word bool 13" : Bool;
      "Alarm Word bool 14" : Bool;
      "Alarm Word bool 15" : Bool;
      "Alarm Word bool 16" : Bool;
      "Delayed Alarm Reset" : TON_TIME;
   END_VAR
BEGIN

REGION Network 1: Check Words